
                               REGION "COPY TO LOCAL"
                                   // remaining time
                                   #elapsedTime := #stations.me[#i].elapsedTime.partReq[#j];
                                   #alottedTime := #stations.me[#i].presetTime.allotted[#j];
                                   #remainingTime := #alottedTime - #elapsedTime;
                                   // critical time
                                   #criticalTime := #stations.me[#i].presetTime.critical[#j];
                               END_REGION

                               REGION "DEFAULT ANIMATION STATE"
                                   IF #remainingTime > #criticalTime THEN
                                       #animation := #anRequested;
                                   END_IF;
                               END_REGION

                               REGION "ORDERED"
                                   IF #partOrdered THEN
                                       #animation := #anPartOrdered;
                                   END_IF;
                               END_REGION

                               REGION "SOLID RED ANIMATION STATE"
                                   IF #remainingTime <= #criticalTime AND #elapsedTime > 0.0 THEN
                                       #animation := #anSolidRed;
                                   END_IF;
                               END_REGION

                               REGION "FLASHING RED ANIMATION STATE
                                   IF #remainingTime <= 0.0 THEN
                                       #animation := #anFlashRed;
                                   END_IF;
                               END_REGION

                           END_IF;
                       END_REGION

                       REGION "PART NOT REQUESTED"
                           IF NOT #partRequested THEN
                               #animation := #anDefault;
                           END_IF;
                       END_REGION

                       REGION "OUTPUT"
                           #stations.me[#i].animations[#j] := #animation;
                       END_REGION

                   END_REGION

               END_FOR;
           END_REGION

       END_FOR;
   END_REGION
END_FUNCTION_BLOCK

FUNCTION_BLOCK "Format Part Call Requests"   // FB9, SCL
{ S7_Optimized_Access := 'TRUE' }
VERSION : 0.1
   VAR_IN_OUT
      requests : "Part Request Data";
      stations : "Stations";
   END_VAR
   VAR
      station : Int;
      button : Int;
   END_VAR
   VAR_TEMP
      address : Int;
      animate : USInt;
      maxRows : Int;
      timeAsReal : Real;
      timeAsTime : WString;
      i : Int;
      inStrRslt : Int;
      invisible : USInt;
      genericVisible : USInt;
      gray : USInt;
      darkGray : USInt;
      red : USInt;
      blue : USInt;
      redFlashing : USInt;
   END_VAR
   VAR CONSTANT
      visible : USInt := 1;
      anDefault : USInt := 0;
      anRequested : USInt := 1;
      anSolidRed : USInt := 2;
      anFlashRed : USInt := 3;
      anPartOrdered : USInt := 4;
   END_VAR
BEGIN
   REGION "COPY TO LOCAL"
       #invisible := "invisible";
       #maxRows := "partReqHmiRowCount";
       #gray := "BgGray";
       #darkGray := "disabled";
       #blue := "BgLBl";
       #red := "BgDRd";
       #redFlashing := "FlDrd";
   END_REGION


   REGION "ITERATE THROUGH VISIBLE TABLE ROWS"
       FOR #i := 0 TO #maxRows DO

           REGION "COPY TO LOCAL"
               #address := UINT_TO_INT(#requests.row[#i].address);
           END_REGION

           REGION "HIDE UNPOPULATED ROWS"
               IF #address = 0 THEN
                   #requests.row[#i].pbSelection.animate := #invisible;
                   #requests.row[#i].rtBackground.animate := #invisible;
                   #animate := 0;
                   #requests.row[#i].tfDropZone.animate := #invisible;
                   #requests.row[#i].tfLine.animate := #invisible;
                   #requests.row[#i].tfPartNumber.animateSL := #invisible;
                   #requests.row[#i].tfPartNumber.animateDL := #invisible;
                   #requests.row[#i].tfTime.animate := #invisible;
               END_IF;
           END_REGION

           REGION "ANIMATE POPULATED ROWS"

               REGION "ANIMATE ROWS WITH DATA"
                   IF #address <> 0 THEN

                       REGION "GET POINTERS FOR STATION ARRAY"
                           #station := #address / 10 - 1;
                           #button := #address MOD 10 - 1;
                       END_REGION

                       REGION "SET ANIMATE"
                           CASE #stations.me[#station].animations[#button] OF
                               #anRequested:
                                   #animate := #gray;
                               #anSolidRed:
                                   #animate := #red;
                               #anFlashRed:
                                   #animate := #redFlashing;
                               #anPartOrdered:
                                   #animate := #blue;
                               ELSE
                                   #animate := #invisible;
                           END_CASE;
                       END_REGION


                       REGION "ANIMATIONS"

                           REGION "PUSHBUTTON VISIBILITY"
                               #requests.row[#i].pbSelection.animate := #visible;
                           END_REGION

                           REGION "BACKGROUND VISIBILITY"
                               #requests.row[#i].rtBackground.animate := #darkGray;
                           END_REGION

                           REGION "DROP ZONE" 
                               #requests.row[#i].tfDropZone.animate := #animate;
                               #requests.row[#i].tfDropZone.value := "Strip Sign"(UINT_TO_WSTRING(#stations.me[#station].dropZone));
                           END_REGION

                           REGION "LINE"
                               #requests.row[#i].tfLine.animate := #animate;
                               #requests.row[#i].tfLine.value := #stations.me[#station].line;
                           END_REGION

                           REGION "PART NUMBER"
                               #requests.row[#i].tfPartNumber.animateSL := #animate;
                               #requests.row[#i].tfPartNumber.value := #stations.me[#station].partNumbers[#button];
                               REGION "DETERMINE VISIBLE ROWS"

                                   REGION "FIND CARRIAGE RETURN"
                                       #inStrRslt := FIND(IN1 := #requests.row[#i].tfPartNumber.value,
                                                          IN2 := wstring#'$L');
                                   END_REGION

                                   REGION "SINGLE LINE"
                                       IF #inStrRslt = 0 THEN
                                           #requests.row[#i].tfPartNumber.animateSL := #animate;
                                           #requests.row[#i].tfPartNumber.animateDL := #invisible;
                                       END_IF;
                                   END_REGION

                                   REGION "DOUBLE LINE"
                                       IF #inStrRslt <> 0 THEN
                                           #requests.row[#i].tfPartNumber.animateSL := #invisible;
                                           #requests.row[#i].tfPartNumber.animateDL := #animate;
                                       END_IF;
                                   END_REGION

                               END_REGION

                           END_REGION

                           REGION "TIME"
                               #requests.row[#i].tfTime.animate := #animate;
                               #timeAsReal := #stations.me[#station].presetTime.allotted[#button];
                               #timeAsReal -= #stations.me[#station].elapsedTime.partReq[#button];
                               #requests.row[#i].tfTime.value := "Real to WString Timer"(#timeAsReal);
                           END_REGION

                       END_REGION

                   END_IF;
               END_REGION

           END_REGION

       END_FOR;
   END_REGION
END_FUNCTION_BLOCK

FUNCTION_BLOCK "KP8 Expanded Animations"   // FB10, SCL
{ S7_Optimized_Access := 'TRUE' }
VERSION : 0.1
   VAR_IN_OUT
      stations : "Stations";
   END_VAR
   VAR_TEMP
      i : Int;
      j : Int;
      colorBox : DWord;
      animation : Int;
      mask : DWord;
   END_VAR
   VAR CONSTANT
      stationCount : Int := 23;
      buttonCount : Int := 7;
      anSolidRed : USInt := 2;
      anFlashRed : USInt := 3;
      anBlue : USInt := 4;
   END_VAR
BEGIN
   REGION "LOOP THROUGH STATIONS"
       FOR #i := 0 TO #stationCount DO

           REGION "LOOP THROUGH BUTTONS"
               FOR #j := 0 TO #buttonCount DO

                   REGION "GET ANIMATION"
                       #animation := #stations.me[#i].animations[#j];
                   END_REGION

                   REGION "SOLID RED"
                       IF #animation = #anSolidRed THEN
                           #colorBox := #stations.me[#i].kp8Out;
                           #mask := 16#FEFEFEFF;
                           #mask := ROL_DWORD(IN := #mask,
                                                 N := INT_TO_UINT(#j));
                           #colorBox := #colorBox AND #mask;
                           #mask := 16#100_0000;
                           #mask := ROL_DWORD(IN := #mask,
                                                 N := INT_TO_UINT(#j));
                           #colorBox := #colorBox OR #mask;
                           #stations.me[#i].kp8Out := #colorBox;
                       END_IF;
                   END_REGION

                   REGION "FLASHING RED"
                       IF #animation = #anFlashRed THEN

                           REGION "RED ON"
                               IF "Clock_1Hz" THEN
                                   #colorBox := #stations.me[#i].kp8Out;
                                   #mask := 16#FEFEFEFF;
                                   #mask := ROL_DWORD(IN := #mask,
                                                         N := INT_TO_UINT(#j));
                                   #colorBox := #colorBox AND #mask;
                                   #mask := 16#100_0000;
                                   #mask := ROL_DWORD(IN := #mask,
                                                         N := INT_TO_UINT(#j));
                                   #colorBox := #colorBox OR #mask;
                                   #stations.me[#i].kp8Out := #colorBox;
                               END_IF;
                           END_REGION

                           REGION "RED OFF"
                               IF NOT "Clock_1Hz" THEN
                                   #colorBox := #stations.me[#i].kp8Out;
                                   #mask := 16#FEFEFEFF;
                                   #mask := ROL_DWORD(IN := #mask,
                                                         N := INT_TO_UINT(#j));
                                   #colorBox := #colorBox AND #mask;
                                   #stations.me[#i].kp8Out := #colorBox;
                               END_IF;
                           END_REGION

                       END_IF;
                   END_REGION

                   REGION "BLUE"
                       IF #animation = #anBlue THEN
                           #colorBox := #stations.me[#i].kp8Out;
                           #mask := 16#FEFEFEFF;
                           #mask := ROL_DWORD(IN := #mask,
                                              N := INT_TO_UINT(#j));
                           #colorBox := #colorBox AND #mask;
                           #mask := 16#0000_0100;
                           #mask := ROL_DWORD(IN := #mask,
                                                 N := INT_TO_UINT(#j));
                           #colorBox := #colorBox OR #mask;
                           #stations.me[#i].kp8Out := #colorBox;
                       END_IF;
                   END_REGION

               END_FOR;
           END_REGION

       END_FOR;
   END_REGION
END_FUNCTION_BLOCK

FUNCTION_BLOCK "Stack Light Animations"   // FB11, SCL
{ S7_Optimized_Access := 'TRUE' }
VERSION : 0.1
   VAR_IN_OUT
      stations : "Stations";
   END_VAR
   VAR_TEMP
      animation : Int;
      i : Int;
      j : Int;
      stackLight : DWord;
   END_VAR
   VAR CONSTANT
      anDefault : USInt := 0;
      anRequested : USInt := 1;
      anSolidRed : USInt := 2;
      anFlashRed : USInt := 3;
      anPartOrdered : USInt := 4;
      buttonCount : Int := 7;
      "Part 01" : Int := 7;
      "Part 01 Green On" : DWord := 16#0400_0000;
      "Part 01 Red On" : DWord := 16#0100_0000;
      "Part 01 Yellow On" : DWord := 16#0200_0000;
      "Part 02" : Int := 3;
      "Part 02 Green On" : DWord := 16#2000_0000;
      "Part 02 Red On" : DWord := 16#0800_0000;
      "Part 02 Yellow On" : DWord := 16#1000_0000;
      "Part 03" : Int := 6;
      "Part 03 Green On" : DWord := 16#0001_0000;
      "Part 03 Red On" : DWord := 16#4000_0000;
      "Part 03 Yellow On" : DWord := 16#8000_0000;
      "Part 04" : Int := 2;
      "Part 04 Green On" : DWord := 16#0008_0000;
      "Part 04 Yellow On" : DWord := 16#0004_0000;
      "Part 04 Red On" : DWord := 16#0002_0000;
      "Part 05" : Int := 5;
      "Part 05 Green On" : DWord := 16#0040_0000;
      "Part 05 Red On" : DWord := 16#0010_0000;
      "Part 05 Yellow On" : DWord := 16#0020_0000;
      "Part 06" : Int := 1;
      "Part 06 Green On" : DWord := 16#0000_0200;
      "Part 06 Red On" : DWord := 16#0080_0000;
      "Part 06 Yellow On" : DWord := 16#0000_0100;
      stationCount : Int := 23;
   END_VAR
BEGIN
   REGION "LOOP THROUGH STATIONS"
       FOR #i := 0 TO #stationCount DO

           REGION "LOOP THROUGH BUTTONS"
               FOR #j := 0 TO #buttonCount DO

                   REGION "COPY INTO LOCAL"
                       #stackLight := #stations.me[#i].stackLightOut;
                       #animation := #stations.me[#i].animations[#j];
                   END_REGION

                   REGION "GREEN"
                       IF #animation = #anDefault THEN
                           CASE #j OF
                               #"Part 01":
                                   #stackLight := #stackLight AND (NOT #"Part 01 Red On");
                                   #stackLight := #stackLight AND (NOT #"Part 01 Yellow On");
                                   #stackLight := #stackLight OR #"Part 01 Green On";
                               #"Part 02":
                                   #stackLight := #stackLight AND (NOT #"Part 02 Red On");
                                   #stackLight := #stackLight AND (NOT #"Part 02 Yellow On");
                                   #stackLight := #stackLight OR #"Part 02 Green On";
                               #"Part 03":
                                   #stackLight := #stackLight AND (NOT #"Part 03 Red On");
                                   #stackLight := #stackLight AND (NOT #"Part 03 Yellow On");
                                   #stackLight := #stackLight OR #"Part 03 Green On";
                               #"Part 04":
                                   #stackLight := #stackLight AND (NOT #"Part 04 Red On");
                                   #stackLight := #stackLight AND (NOT #"Part 04 Yellow On");
                                   #stackLight := #stackLight OR #"Part 04 Green On";
                               #"Part 05":
                                   #stackLight := #stackLight AND (NOT #"Part 05 Red On");
                                   #stackLight := #stackLight AND (NOT #"Part 05 Yellow On");
                                   #stackLight := #stackLight OR #"Part 05 Green On";
                               #"Part 06":
                                   #stackLight := #stackLight AND (NOT #"Part 06 Red On");
                                   #stackLight := #stackLight AND (NOT #"Part 06 Yellow On");
                                   #stackLight := #stackLight OR #"Part 06 Green On";
                               ELSE
                                   ;
                           END_CASE;
                       END_IF;
                   END_REGION

                   REGION "YELLOW"
                       IF #animation = #anRequested THEN
                           CASE #j OF
                               #"Part 01":
                                   #stackLight := #stackLight AND (NOT #"Part 01 Red On");
                                   #stackLight := #stackLight OR #"Part 01 Yellow On";
                                   #stackLight := #stackLight AND (NOT #"Part 01 Green On");
                               #"Part 02":
                                   #stackLight := #stackLight AND (NOT #"Part 02 Red On");
                                   #stackLight := #stackLight OR #"Part 02 Yellow On";
                                   #stackLight := #stackLight AND (NOT #"Part 02 Green On");
                               #"Part 03":
                                   #stackLight := #stackLight AND (NOT #"Part 03 Red On");
                                   #stackLight := #stackLight OR #"Part 03 Yellow On";
                                   #stackLight := #stackLight AND (NOT #"Part 03 Green On");
                               #"Part 04":
                                   #stackLight := #stackLight AND (NOT #"Part 04 Red On");
                                   #stackLight := #stackLight OR #"Part 04 Yellow On";
                                   #stackLight := #stackLight AND (NOT #"Part 04 Green On");
                               #"Part 05":
                                   #stackLight := #stackLight AND (NOT #"Part 05 Red On");
                                   #stackLight := #stackLight OR #"Part 05 Yellow On";
                                   #stackLight := #stackLight AND (NOT #"Part 05 Green On");
                               #"Part 06":
                                   #stackLight := #stackLight AND (NOT #"Part 06 Red On");
                                   #stackLight := #stackLight OR #"Part 06 Yellow On";
                                   #stackLight := #stackLight AND (NOT #"Part 06 Green On");
                               ELSE
                                   ;
                           END_CASE;
                       END_IF;
                   END_REGION

                   REGION "SOLID RED"
                       IF #animation = #anSolidRed THEN
                           CASE #j OF
                               #"Part 01":
                                   #stackLight := #stackLight OR #"Part 01 Red On";
                                   #stackLight := #stackLight AND (NOT #"Part 01 Yellow On");
                                   #stackLight := #stackLight AND (NOT #"Part 01 Green On");
                               #"Part 02":
                                   #stackLight := #stackLight OR #"Part 02 Red On";
                                   #stackLight := #stackLight AND (NOT #"Part 02 Yellow On");
                                   #stackLight := #stackLight AND (NOT #"Part 02 Green On");
                               #"Part 03":
                                   #stackLight := #stackLight OR #"Part 03 Red On";
                                   #stackLight := #stackLight AND (NOT #"Part 03 Yellow On");
                                   #stackLight := #stackLight AND (NOT #"Part 03 Green On");
                               #"Part 04":
                                   #stackLight := #stackLight OR #"Part 04 Red On";
                                   #stackLight := #stackLight AND (NOT #"Part 04 Yellow On");
                                   #stackLight := #stackLight AND (NOT #"Part 04 Green On");
                               #"Part 05":
                                   #stackLight := #stackLight OR #"Part 05 Red On";
                                   #stackLight := #stackLight AND (NOT #"Part 05 Yellow On");
                                   #stackLight := #stackLight AND (NOT #"Part 05 Green On");
                               #"Part 06":
                                   #stackLight := #stackLight OR #"Part 06 Red On";
                                   #stackLight := #stackLight AND (NOT #"Part 06 Yellow On");
                                   #stackLight := #stackLight AND (NOT #"Part 06 Green On");
                               ELSE
                                   ;
                           END_CASE;
                       END_IF;
                   END_REGION

                   REGION "FLASHING RED"
                       IF #animation = #anFlashRed THEN

                           REGION "RED ON"
                               IF "Clock_1Hz" THEN
                                   CASE #j OF
                                       #"Part 01":
                                           #stackLight := #stackLight OR #"Part 01 Red On";
                                           #stackLight := #stackLight AND (NOT #"Part 01 Yellow On");
                                           #stackLight := #stackLight AND (NOT #"Part 01 Green On");
                                       #"Part 02":
                                           #stackLight := #stackLight OR #"Part 02 Red On";
                                           #stackLight := #stackLight AND (NOT #"Part 02 Yellow On");
                                           #stackLight := #stackLight AND (NOT #"Part 02 Green On");
                                       #"Part 03":
                                           #stackLight := #stackLight OR #"Part 03 Red On";
                                           #stackLight := #stackLight AND (NOT #"Part 03 Yellow On");
                                           #stackLight := #stackLight AND (NOT #"Part 03 Green On");
                                       #"Part 04":
                                           #stackLight := #stackLight OR #"Part 04 Red On";
                                           #stackLight := #stackLight AND (NOT #"Part 04 Yellow On");
                                           #stackLight := #stackLight AND (NOT #"Part 04 Green On");
                                       #"Part 05":
                                           #stackLight := #stackLight OR #"Part 05 Red On";
                                           #stackLight := #stackLight AND (NOT #"Part 05 Yellow On");
                                           #stackLight := #stackLight AND (NOT #"Part 05 Green On");
                                       #"Part 06":
                                           #stackLight := #stackLight OR #"Part 06 Red On";
                                           #stackLight := #stackLight AND (NOT #"Part 06 Yellow On");
                                           #stackLight := #stackLight AND (NOT #"Part 06 Green On");
                                       ELSE
                                           ;
                                   END_CASE;
                               END_IF;
                           END_REGION

                           REGION "RED OFF"
                               IF NOT "Clock_1Hz" THEN
                                   CASE #j OF
                                       #"Part 01":
                                           #stackLight := #stackLight AND (NOT #"Part 01 Red On");
                                           #stackLight := #stackLight AND (NOT #"Part 01 Yellow On");
                                           #stackLight := #stackLight AND (NOT #"Part 01 Green On");
                                       #"Part 02":
                                           #stackLight := #stackLight AND (NOT #"Part 02 Red On");
                                           #stackLight := #stackLight AND (NOT #"Part 02 Yellow On");
                                           #stackLight := #stackLight AND (NOT #"Part 02 Green On");
                                       #"Part 03":
                                           #stackLight := #stackLight AND (NOT #"Part 03 Red On");
                                           #stackLight := #stackLight AND (NOT #"Part 03 Yellow On");
                                           #stackLight := #stackLight AND (NOT #"Part 03 Green On");
                                       #"Part 04":
                                           #stackLight := #stackLight AND (NOT #"Part 04 Red On");
                                           #stackLight := #stackLight AND (NOT #"Part 04 Yellow On");
                                           #stackLight := #stackLight AND (NOT #"Part 04 Green On");
                                       #"Part 05":
                                           #stackLight := #stackLight AND (NOT #"Part 05 Red On");
                                           #stackLight := #stackLight AND (NOT #"Part 05 Yellow On");
                                           #stackLight := #stackLight AND (NOT #"Part 05 Green On");
                                       #"Part 06":
                                           #stackLight := #stackLight AND (NOT #"Part 06 Red On");
                                           #stackLight := #stackLight AND (NOT #"Part 06 Yellow On");
                                           #stackLight := #stackLight AND (NOT #"Part 06 Green On");
                                       ELSE
                                           ;
                                   END_CASE;
                               END_IF;
                           END_REGION

                       END_IF;
                   END_REGION

                   REGION "COPY OUT TO GLOBAL"
                       #stations.me[#i].stackLightOut := #stackLight;
                   END_REGION

               END_FOR;
           END_REGION

       END_FOR;
   END_REGION
END_FUNCTION_BLOCK

FUNCTION_BLOCK "KP8 Button Activation"   // FB12, SCL
{ S7_Optimized_Access := 'TRUE' }
VERSION : 0.1
   VAR_IN_OUT
      stations : "Stations";
   END_VAR
   VAR
      old : Struct
         kp8Config : Array[0.."stnCount"] of "KP8 Button Config";
      END_STRUCT;
   END_VAR
   VAR_TEMP
      btnCount : Int;
      currentPNs : Array[0..7] of WString[40];
      i : Int;
      init : Bool;
      j : Int;
      stnCount : Int;
      temp : Int;
   END_VAR
BEGIN
   REGION "GET STATION COUNT"
       #stnCount := "stnCount";
       #btnCount := "ptsPerStn";
   END_REGION

   REGION "LOOP THROUGH STATIONS"
       FOR #i := 0 TO #stnCount DO

           REGION "COPY TO LOCAL"
               #currentPNs := #stations.me[#i].partNumbers;
           END_REGION


           REGION "LOOP THROUGH BUTTONS"
               FOR #j := 0 TO #btnCount DO

                       REGION "ACTIVATE BUTTON"
                           IF LEN(#currentPNs[#j]) <> 0 THEN
                               #stations.me[#i].kp8Config.activate[#j] := TRUE;
                               #stations.me[#i].kp8Config.colorOff[#j] := 'green';
                               #stations.me[#i].kp8Config.colorOn1[#j] := 'yellow';
                               #stations.me[#i].kp8Config.colorOn2[#j] := '';
                               #stations.me[#i].kp8Config.flash[#j] := FALSE;
                               #stations.me[#i].kp8Config.group[#j] := 0;
                               #stations.me[#i].kp8Config.mode[#j] := TRUE;
                           END_IF;
                       END_REGION

                       REGION "DEACTIVATE BUTTON"
                           IF LEN(#currentPNs[#j]) = 0 THEN
                               #stations.me[#i].kp8Config.activate[#j] := FALSE;
                               #stations.me[#i].kp8Config.colorOff[#j] := '';
                               #stations.me[#i].kp8Config.colorOn1[#j] := '';
                               #stations.me[#i].kp8Config.colorOn2[#j] := '';
                               #stations.me[#i].kp8Config.flash[#j] := FALSE;
                               #stations.me[#i].kp8Config.group[#j] := 0;
                               #stations.me[#i].kp8Config.mode[#j] := FALSE;
                           END_IF;
                       END_REGION

               END_FOR;
           END_REGION

           REGION "SOFT INIT"
               IF #stations.me[#i].kp8Config <> #old.kp8Config[#i] THEN
                   #stations.me[#i].init.soft := TRUE;
               END_IF;
           END_REGION

           REGION "SAVE FOR CHANGE DETECTION"
               #old.kp8Config[#i] := #stations.me[#i].kp8Config;
           END_REGION

       END_FOR;
   END_REGION
END_FUNCTION_BLOCK

FUNCTION_BLOCK "Remove Part Request"   // FB13, SCL
{ S7_Optimized_Access := 'TRUE' }
VERSION : 0.1
   VAR_IN_OUT
      pRow : Int;
      requests : "Part Request Data";
      stations : "Stations";
   END_VAR
   VAR
      old : Struct
         partReq : "Station Old Presses";
      END_STRUCT;
   END_VAR
   VAR_TEMP
      address : UInt;
      blankRow : "Table Row";
      hasPart : Bool;
      i : Int;
      j : Int;
      k : Int;
      logAddress : UInt;
      maxRows : Int;
      noPart : Bool;
      oldPartReq : Bool;
      partNumber : WString;
      partReq : Bool;
      pRemoveRow : Int;
      btnCount : Int;
      stnCount : Int;
      removeAddress : Bool;
   END_VAR
BEGIN
   REGION "COPY TO LOCAL"
       #maxRows := "partReqHmiRowCount";
       #stnCount := "stnCount";
       #btnCount := "ptsPerStn";
   END_REGION


   REGION "FOR EACH STATION"
       FOR #i := 0 TO #stnCount DO

           REGION "FOR EACH BUTTON"
               FOR #j := 1 TO #btnCount DO

                   REGION "COPY TO LOCAL"
                       #partReq := #stations.me[#i].btnStates[#j];
                       #oldPartReq := #old.partReq.me[#i, #j];
                   END_REGION

                   REGION "DETERMINE STATE"

                       REGION "PART REQUEST FALLING EDGE"
                           IF NOT #partReq AND #oldPartReq THEN

                               REGION "SAVE FOR CHANGE DETECTION"
                                   #old.partReq.me[#i, #j] := #partReq;
                               END_REGION

                               REGION "COPY TO LOCAL"
                                   #partNumber := #stations.me[#i].partNumbers[#j];
                               END_REGION

                               REGION "BUTTON HAS NO PART"
                                   IF #partNumber = wstring#'' THEN
                                       #hasPart := FALSE;
                                       #noPart := TRUE;
                                   END_IF;
                               END_REGION

                               REGION "BUTTON HAS PART"
                                   IF #partNumber <> wstring#'' THEN
                                       #hasPart := TRUE;
                                       #noPart := FALSE;
                                   END_IF;
                               END_REGION

                           END_IF;
                       END_REGION

                   END_REGION

                   REGION "NO PART"
                       IF #noPart THEN

                           REGION "TURN OFF THE LIGHTS"
                               #hasPart := FALSE;
                               #noPart := FALSE;
                           END_REGION

                       END_IF;

                   END_REGION

                   REGION "HAS PART"
                       IF #hasPart THEN

                           REGION "TURN OFF THE LIGHTS"
                               #hasPart := FALSE;
                           END_REGION

                           REGION "CALCULATE ADDRESS"
                               #address := (INT_TO_UINT(#i) + 1) * 10 + (INT_TO_UINT(#j) + 1);
                           END_REGION

                           REGION "RESET FLAG"
                               #removeAddress := FALSE;
                           END_REGION

                           REGION "SEARCH EACH ROW IN PART DB"
                               FOR #k := 0 TO #maxRows DO

                                   REGION "COPY TO LOCAL"
                                       #logAddress := #requests.row[#k].address;
                                   END_REGION

                                   REGION "ON MATCH"
                                       IF #logAddress = #address THEN

                                           REGION "SET FLAG"
                                               #removeAddress := TRUE;
                                           END_REGION

                                           REGION "SAVE POINTER"
                                               #pRemoveRow := #k;
                                           END_REGION

                                       END_IF;
                                   END_REGION

                               END_FOR;
                           END_REGION

                       END_IF;
                   END_REGION

                   REGION "REMOVE ADDRESS"
                       IF #removeAddress THEN

                           REGION "TURN OFF THE LIGHTS"
                               #removeAddress := FALSE;
                           END_REGION

                           REGION "TURN OFF REQUEST"
                               #stations.me[#i].partRequested[#j] := FALSE;
                           END_REGION

                           REGION "REMOVAL PROCESS"

                               REGION "REMOVE ROW"
                                   #requests.row[#pRemoveRow] := #blankRow;
                               END_REGION

                               REGION "REMOVE PART ORDERED"
                                   #stations.me[#i].partOrdered[#j] := FALSE;
                               END_REGION

                           END_REGION

                           REGION "ROW POINTER"

                               REGION "DECREMENT"
                                   #pRow := #pRow - 1;
                               END_REGION

                               REGION "LOW LIMIT ROLL OVER"
                                   IF #pRow < 0 THEN
                                       #pRow := 0;
                                   END_IF;
                               END_REGION

                           END_REGION

                       END_IF;
                   END_REGION

               END_FOR;

           END_REGION

       END_FOR;
   END_REGION
END_FUNCTION_BLOCK

FUNCTION_BLOCK "HMI Settings Screen"   // FB14, LAD
{ S7_Optimized_Access := 'TRUE' }
VERSION : 0.1
   VAR_IN_OUT
      settings : "Settings";
      stations : "Stations";
   END_VAR
   VAR
      tmrTimeOut : TON_TIME;
      instStaSel : "Station Selection";
      instKP8BtnSel : "KP8 Button Selections";
      old : Struct
         asgnPN : Bool;
         asgnAlloted : Bool;
         asgnCritical : Bool;
         nextPress : Bool;
         prevPress : Bool;
         selBtnCount : Int;
         selBtnNumber : Int;
         selStnCount : Int;
         selStnNumber : Int;
      END_STRUCT;
      instAsnBtnPrms : "Assign Button Parameters";
      instAniPNTmr : "Animate: PN & Timers";
   END_VAR
   VAR_TEMP
      pBN : Int;
      pSN : Int;
      wStringBox : WString;
   END_VAR
   VAR CONSTANT
      ptTimeOut : Time := t#15m;
   END_VAR
   VAR_TEMP   // added for the SCL form of the ladder/FBD networks
      _w1 : Bool;
   END_VAR
BEGIN

REGION Network 1: ENTRY TIMEOUT
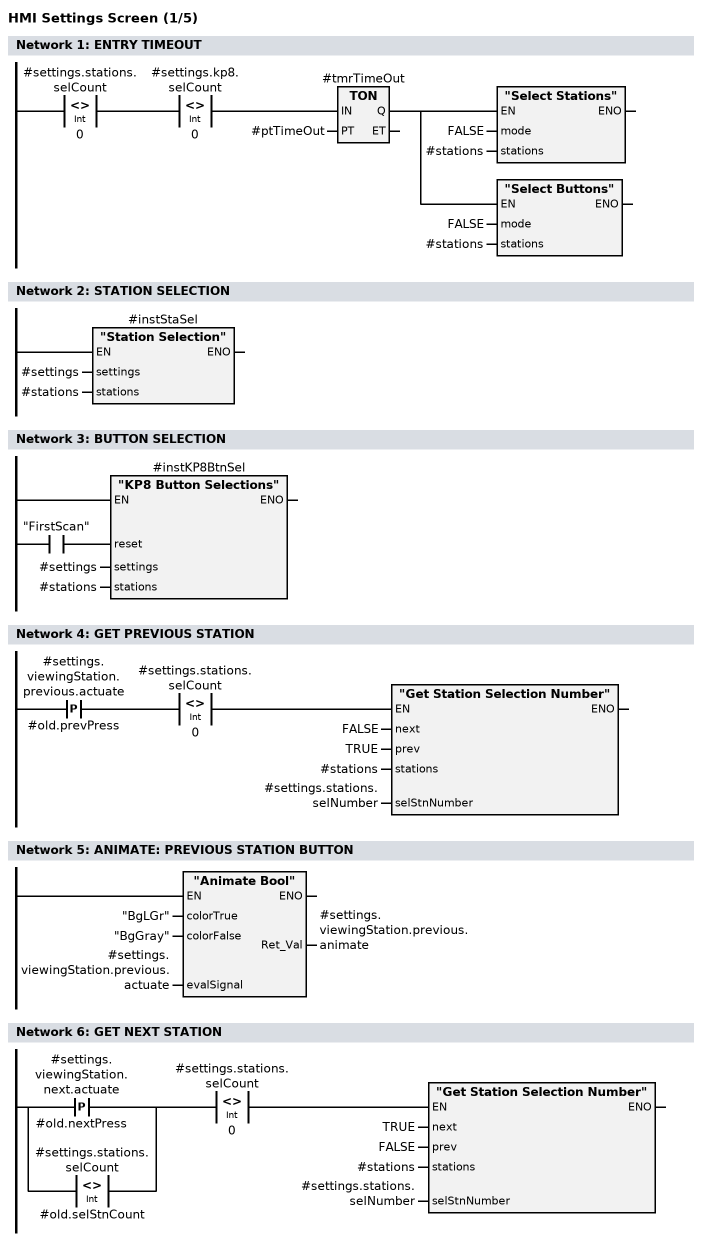
   #tmrTimeOut(IN := (#settings.stations.selCount <> 0) AND (#settings.kp8.selCount <> 0), PT := #ptTimeOut);   // TON
   IF #tmrTimeOut.Q THEN
       "Select Stations"(mode := FALSE, stations := #stations);
       "Select Buttons"(mode := FALSE, stations := #stations);
   END_IF;
END_REGION

REGION Network 2: STATION SELECTION
   RUNG wire#powerrail
      #instStaSel(settings := #settings, stations := #stations)
   END_RUNG
   // the same network as SCL:
   #instStaSel(settings := #settings, stations := #stations);   // "Station Selection"
END_REGION

REGION Network 3: BUTTON SELECTION
   RUNG wire#powerrail
      #instKP8BtnSel(reset := wire#w1, settings := #settings, stations := #stations)
   END_RUNG
   RUNG wire#powerrail
      Contact( "FirstScan" )
   END_RUNG wire#w1
   // the same network as SCL:
   #instKP8BtnSel(reset := "FirstScan", settings := #settings, stations := #stations);   // "KP8 Button Selections"
END_REGION

REGION Network 4: GET PREVIOUS STATION
   RUNG wire#powerrail
      P_Contact(operand := #settings.viewingStation.previous.actuate, bit := #old.prevPress)
      { S7_Templates := "SrcType := Int" } NE_Contact(in1 := #settings.stations.selCount, in2 := 0)
      "Get Station Selection Number"(next := FALSE, prev := TRUE, stations := #stations, selStnNumber := #settings.stations.selNumber)
   END_RUNG
   // the same network as SCL:
   #_w1 := #settings.viewingStation.previous.actuate AND NOT #old.prevPress;   // rising edge of #settings.viewingStation.previous.actuate
   #old.prevPress := #settings.viewingStation.previous.actuate;
   IF #_w1 AND (#settings.stations.selCount <> 0) THEN
       "Get Station Selection Number"(next := FALSE,
                               prev := TRUE,
                               stations := #stations,
                               selStnNumber := #settings.stations.selNumber);
   END_IF;
END_REGION

REGION Network 5: ANIMATE: PREVIOUS STATION BUTTON
   RUNG wire#powerrail
      "Animate Bool"(colorTrue := "BgLGr", colorFalse := "BgGray", evalSignal := #settings.viewingStation.previous.actuate, Ret_Val => #settings.viewingStation.previous.animate)
   END_RUNG
   // the same network as SCL:
   #settings.viewingStation.previous.animate := "Animate Bool"(colorTrue := "BgLGr",
                           colorFalse := "BgGray",
                           evalSignal := #settings.viewingStation.previous.actuate);
END_REGION

REGION Network 6: GET NEXT STATION
   RUNG wire#powerrail
      P_Contact(operand := #settings.viewingStation.next.actuate, bit := #old.nextPress)
      wire#w1
      { S7_Templates := "SrcType := Int" } NE_Contact(in1 := #settings.stations.selCount, in2 := 0)
      "Get Station Selection Number"(next := TRUE, prev := FALSE, stations := #stations, selStnNumber := #settings.stations.selNumber)
   END_RUNG
   RUNG wire#powerrail
      { S7_Templates := "SrcType := Int" } NE_Contact(in1 := #settings.stations.selCount, in2 := #old.selStnCount)
   END_RUNG wire#w1
   // the same network as SCL:
   #_w1 := #settings.viewingStation.next.actuate AND NOT #old.nextPress;   // rising edge of #settings.viewingStation.next.actuate
   #old.nextPress := #settings.viewingStation.next.actuate;
   IF (#_w1 OR (#settings.stations.selCount <> #old.selStnCount)) AND (#settings.stations.selCount <> 0) THEN
       "Get Station Selection Number"(next := TRUE,
                               prev := FALSE,
                               stations := #stations,
                               selStnNumber := #settings.stations.selNumber);
   END_IF;
END_REGION

REGION Network 7: ANIMATE: NEXT STATION BUTTON
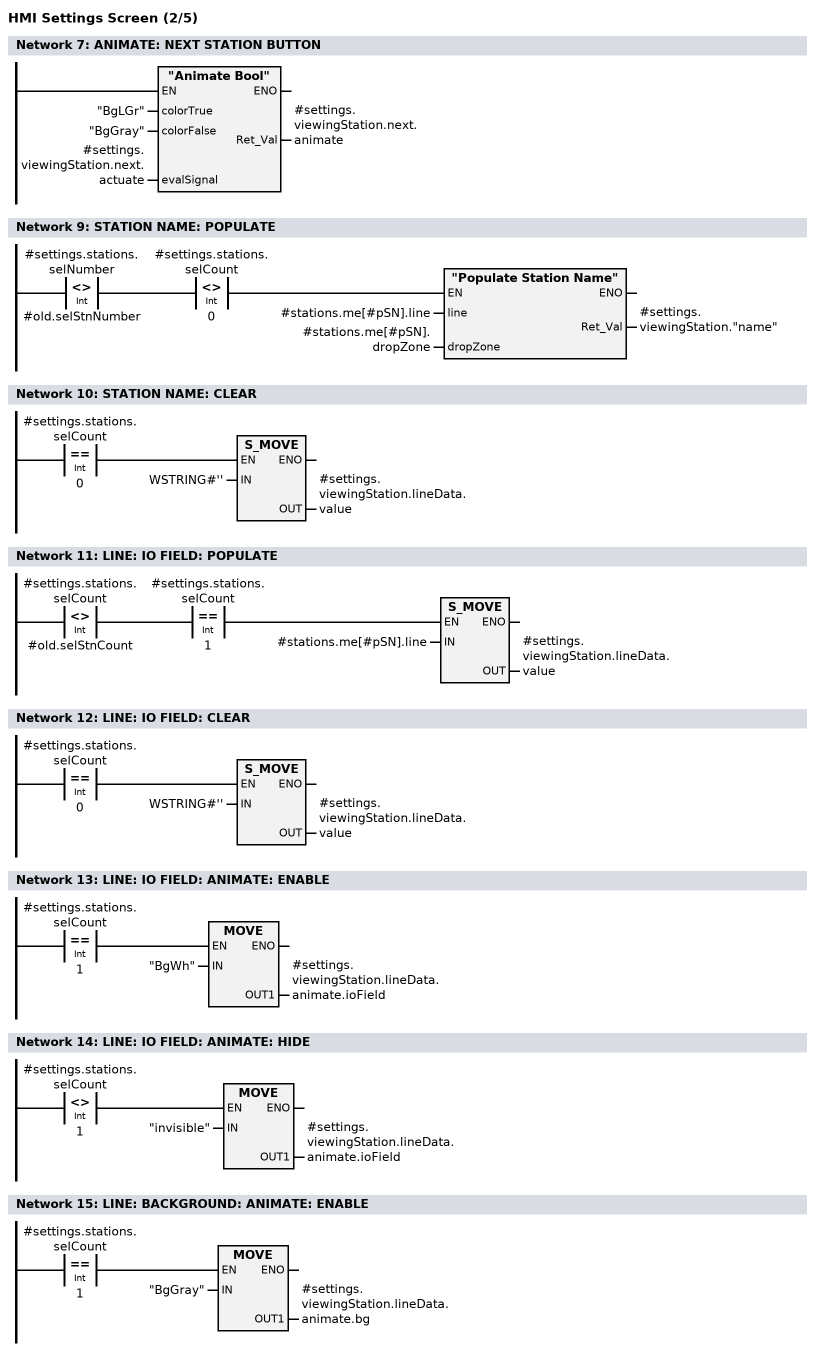
   RUNG wire#powerrail
      "Animate Bool"(colorTrue := "BgLGr", colorFalse := "BgGray", evalSignal := #settings.viewingStation.next.actuate, Ret_Val => #settings.viewingStation.next.animate)
   END_RUNG
   // the same network as SCL:
   #settings.viewingStation.next.animate := "Animate Bool"(colorTrue := "BgLGr",
                           colorFalse := "BgGray",
                           evalSignal := #settings.viewingStation.next.actuate);
END_REGION

REGION Network 8 (SCL): COPY TO POINTERS
   #pSN := #settings.stations.selNumber;
   #pBN := #settings.kp8.selBtnNumber;
END_REGION

REGION Network 9: STATION NAME: POPULATE
   RUNG wire#powerrail
      { S7_Templates := "SrcType := Int" } NE_Contact(in1 := #settings.stations.selNumber, in2 := #old.selStnNumber)
      { S7_Templates := "SrcType := Int" } NE_Contact(in1 := #settings.stations.selCount, in2 := 0)
      "Populate Station Name"(line := #stations.me[#pSN].line, dropZone := #stations.me[#pSN].dropZone, Ret_Val => #settings.viewingStation."name")
   END_RUNG
   // the same network as SCL:
   IF (#settings.stations.selNumber <> #old.selStnNumber) AND (#settings.stations.selCount <> 0) THEN
       #settings.viewingStation."name" := "Populate Station Name"(line := #stations.me[#pSN].line,
                               dropZone := #stations.me[#pSN].dropZone);
   END_IF;
END_REGION

REGION Network 10: STATION NAME: CLEAR
   RUNG wire#powerrail
      { S7_Templates := "SrcType := Int" } EQ_Contact(in1 := #settings.stations.selCount, in2 := 0)
      S_Move(in := WSTRING#'', out => #settings.viewingStation.lineData.value)
   END_RUNG
   // the same network as SCL:
   IF #settings.stations.selCount = 0 THEN #settings.viewingStation.lineData.value := WSTRING#''; END_IF;
END_REGION

REGION Network 11: LINE: IO FIELD: POPULATE
   RUNG wire#powerrail
      { S7_Templates := "SrcType := Int" } NE_Contact(in1 := #settings.stations.selCount, in2 := #old.selStnCount)
      { S7_Templates := "SrcType := Int" } EQ_Contact(in1 := #settings.stations.selCount, in2 := 1)
      S_Move(in := #stations.me[#pSN].line, out => #settings.viewingStation.lineData.value)
   END_RUNG
   // the same network as SCL:
   IF (#settings.stations.selCount <> #old.selStnCount) AND (#settings.stations.selCount = 1) THEN
       #settings.viewingStation.lineData.value := #stations.me[#pSN].line;
   END_IF;
END_REGION

REGION Network 12: LINE: IO FIELD: CLEAR
   RUNG wire#powerrail
      { S7_Templates := "SrcType := Int" } EQ_Contact(in1 := #settings.stations.selCount, in2 := 0)
      S_Move(in := WSTRING#'', out => #settings.viewingStation.lineData.value)
   END_RUNG
   // the same network as SCL:
   IF #settings.stations.selCount = 0 THEN #settings.viewingStation.lineData.value := WSTRING#''; END_IF;
END_REGION

REGION Network 13: LINE: IO FIELD: ANIMATE: ENABLE
   RUNG wire#powerrail
      { S7_Templates := "SrcType := Int" } EQ_Contact(in1 := #settings.stations.selCount, in2 := 1)
      Move(in := "BgWh", out1 => #settings.viewingStation.lineData.animate.ioField)
   END_RUNG
   // the same network as SCL:
   IF #settings.stations.selCount = 1 THEN
       #settings.viewingStation.lineData.animate.ioField := "BgWh";
   END_IF;
END_REGION

REGION Network 14: LINE: IO FIELD: ANIMATE: HIDE
   RUNG wire#powerrail
      { S7_Templates := "SrcType := Int" } NE_Contact(in1 := #settings.stations.selCount, in2 := 1)
      Move(in := "invisible", out1 => #settings.viewingStation.lineData.animate.ioField)
   END_RUNG
   // the same network as SCL:
   IF #settings.stations.selCount <> 1 THEN
       #settings.viewingStation.lineData.animate.ioField := "invisible";
   END_IF;
END_REGION

REGION Network 15: LINE: BACKGROUND: ANIMATE: ENABLE
   RUNG wire#powerrail
      { S7_Templates := "SrcType := Int" } EQ_Contact(in1 := #settings.stations.selCount, in2 := 1)
      Move(in := "BgGray", out1 => #settings.viewingStation.lineData.animate.bg)
   END_RUNG
   // the same network as SCL:
   IF #settings.stations.selCount = 1 THEN #settings.viewingStation.lineData.animate.bg := "BgGray"; END_IF;
END_REGION

REGION Network 16: LINE: BACKGROUND: ANIMATE: HIDE
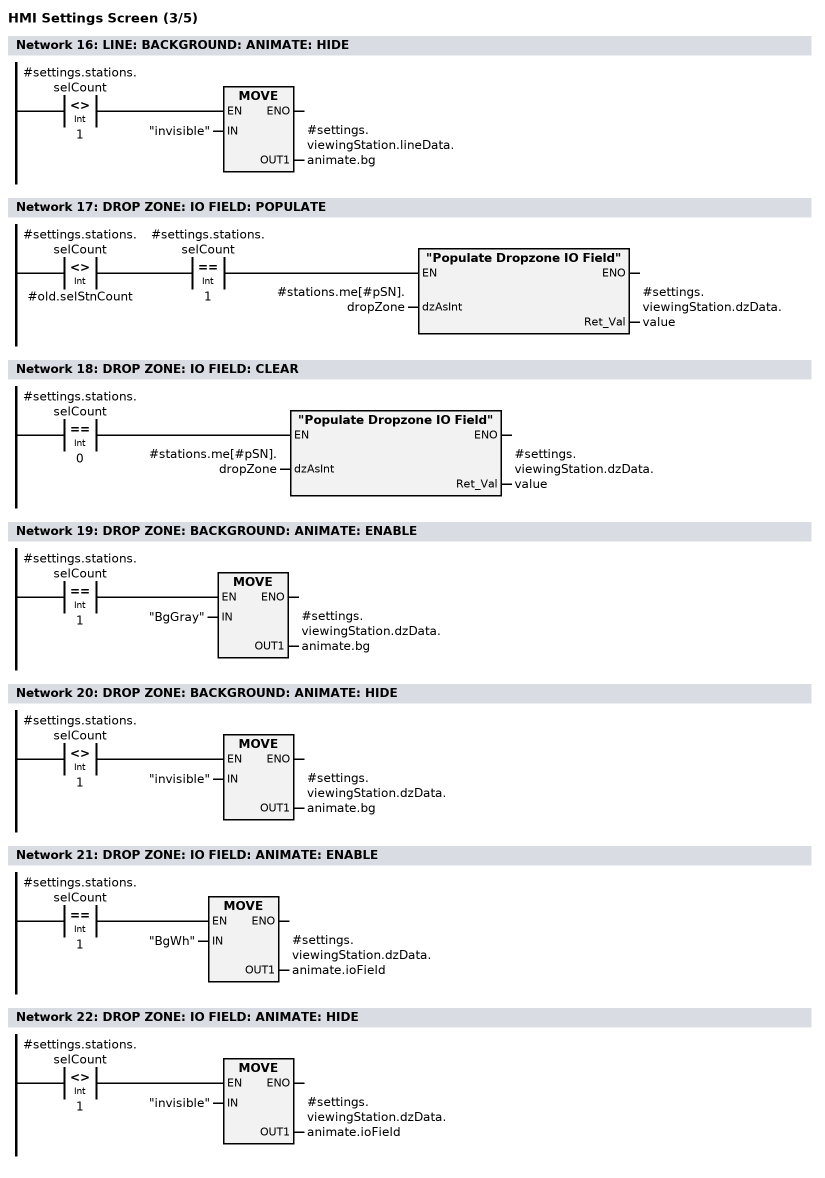
   RUNG wire#powerrail
      { S7_Templates := "SrcType := Int" } NE_Contact(in1 := #settings.stations.selCount, in2 := 1)
      Move(in := "invisible", out1 => #settings.viewingStation.lineData.animate.bg)
   END_RUNG
   // the same network as SCL:
   IF #settings.stations.selCount <> 1 THEN
       #settings.viewingStation.lineData.animate.bg := "invisible";
   END_IF;
END_REGION

REGION Network 17: DROP ZONE: IO FIELD: POPULATE
   RUNG wire#powerrail
      { S7_Templates := "SrcType := Int" } NE_Contact(in1 := #settings.stations.selCount, in2 := #old.selStnCount)
      { S7_Templates := "SrcType := Int" } EQ_Contact(in1 := #settings.stations.selCount, in2 := 1)
      "Populate Dropzone IO Field"(dzAsInt := #stations.me[#pSN].dropZone, Ret_Val => #settings.viewingStation.dzData.value)
   END_RUNG
   // the same network as SCL:
   IF (#settings.stations.selCount <> #old.selStnCount) AND (#settings.stations.selCount = 1) THEN
       #settings.viewingStation.dzData.value := "Populate Dropzone IO Field"(dzAsInt := #stations.me[#pSN].dropZone);
   END_IF;
END_REGION

REGION Network 18: DROP ZONE: IO FIELD: CLEAR
   RUNG wire#powerrail
      { S7_Templates := "SrcType := Int" } EQ_Contact(in1 := #settings.stations.selCount, in2 := 0)
      "Populate Dropzone IO Field"(dzAsInt := #stations.me[#pSN].dropZone, Ret_Val => #settings.viewingStation.dzData.value)
   END_RUNG
   // the same network as SCL:
   IF #settings.stations.selCount = 0 THEN
       #settings.viewingStation.dzData.value := "Populate Dropzone IO Field"(dzAsInt := #stations.me[#pSN].dropZone);
   END_IF;
END_REGION

REGION Network 19: DROP ZONE: BACKGROUND: ANIMATE: ENABLE
   RUNG wire#powerrail
      { S7_Templates := "SrcType := Int" } EQ_Contact(in1 := #settings.stations.selCount, in2 := 1)
      Move(in := "BgGray", out1 => #settings.viewingStation.dzData.animate.bg)
   END_RUNG
   // the same network as SCL:
   IF #settings.stations.selCount = 1 THEN #settings.viewingStation.dzData.animate.bg := "BgGray"; END_IF;
END_REGION

REGION Network 20: DROP ZONE: BACKGROUND: ANIMATE: HIDE
   RUNG wire#powerrail
      { S7_Templates := "SrcType := Int" } NE_Contact(in1 := #settings.stations.selCount, in2 := 1)
      Move(in := "invisible", out1 => #settings.viewingStation.dzData.animate.bg)
   END_RUNG
   // the same network as SCL:
   IF #settings.stations.selCount <> 1 THEN
       #settings.viewingStation.dzData.animate.bg := "invisible";
   END_IF;
END_REGION

